(* Logix 5000 project; controller MV vendor 1 type 14 code 217 rev 31.11; software revision 31.00; part 24 of 53 *)
(* tags used below, declared in another part *)
   CheckTimeMask : INT;
   CWD : CHECKWORD_FLAGS;
   Delphi_Does_Eng_Func : BOOL;
   MC_CH1_FM_AI : PlantItem;   // CH1_FM
   MC_CH1_PTX_AI : PlantItem;   // CH1_PTX
   MC_CH2_FM_AI : PlantItem;   // CH2_FM
   MC_CH2_PTX_AI : PlantItem;   // CH2_PTX
   MC_CIP_AV09 : PlantItem;   // CIP_AV09
   MC_N100 : INT[255];   // C1_PLC Channel 1 PLC data
   MC_N100_29_1_Storagebit : BOOL;
   MC_N100_29_2_Storagebit : BOOL;
   MC_N100_29_3_Storagebit : BOOL;
   MC_N100_29_4_Storagebit : BOOL;
   MC_N102 : INT[255];   // CH1 PROG Channel 1 CIP progra m
   MC_N120 : INT[255];   // C2 PLC Channel 2 PLC data
   MC_N120_29_1_Storagebit : BOOL;
   MC_N120_29_2_Storagebit : BOOL;
   MC_N120_29_3_Storagebit : BOOL;
   MC_N120_29_4_Storagebit : BOOL;
   MC_N122 : INT[255];   // CH2 PROG Channel 2 CIP progra m
   MC_N20 : INT[255];   // P1 PRESS Control block and da ta for P1 pressure P ID loop
   MC_N21 : INT[255];   // P1 FLOW Control block and da ta for P1 flowrate P ID loop
   MC_N22 : INT[255];   // P2 PRESS Control block and da ta for P2 pressure P ID loop
   MC_N23 : INT[255];   // P2 FLOW Control block and da ta for P2 flowrate P ID loop
   MC_N255 : INT[255];   // CHECKWORDS Plant item checkword s
   MC_P1 : PlantItem;   // P1
   MC_P1_Flow_PID : PID;
   MC_P1_Flow_PID_Output : REAL;
   MC_P1_Pressure_PID : PID;
   MC_P1_Pressure_PID_Output : REAL;
   MC_P1_SP_AO : PlantItem;   // P1_SP
   MC_P2 : PlantItem;   // P2
   MC_P2_Flow_PID : PID;
   MC_P2_Flow_PID_Output : REAL;
   MC_P2_Pressure_PID : PID;
   MC_P2_Pressure_PID_Output : REAL;
   MC_P2_SP_AO : PlantItem;   // P2_SP
   TempChecktime : DINT;
(* MC_Common, continued *)

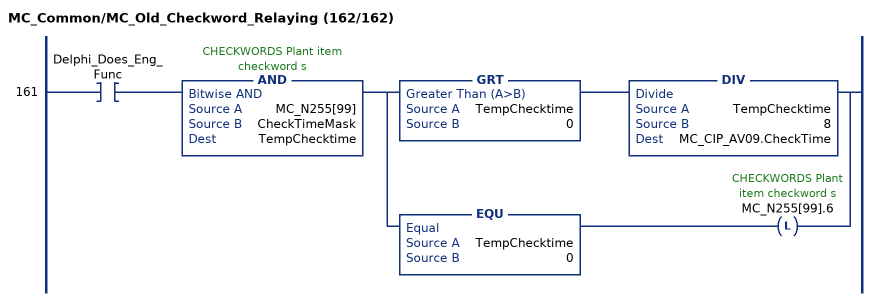
   [picture p434: MC_Common/MC_Old_Checkword_Relaying rungs 161-161]
   161: XIC(Delphi_Does_Eng_Func)AND(MC_N255[99],CheckTimeMask,TempChecktime)[GRT(TempChecktime,0) DIV(TempChecktime,8,MC_CIP_AV09.CheckTime) ,EQU(TempChecktime,0) OTL(MC_N255[99].6) ];
END_ROUTINE

ROUTINE MC_P1_FLOW_21   (* ladder *)
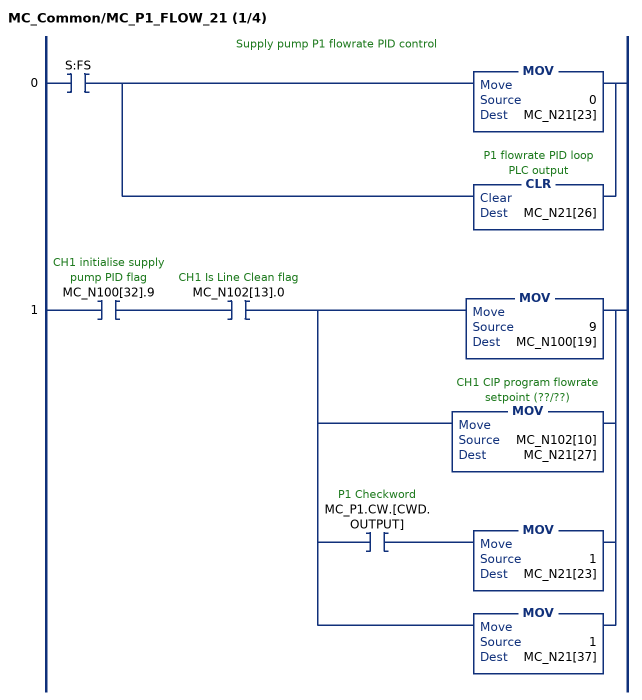
   // Supply pump P1 flowrate PID control
   0: XIC(S:FS)[MOV(0,MC_N21[23]) ,CLR(MC_N21[26]) ];
   1: XIC(MC_N100[32].9)XIC(MC_N102[13].0)[MOV(9,MC_N100[19]) ,MOV(MC_N102[10],MC_N21[27]) ,XIC(MC_P1.CW.[CWD.OUTPUT]) MOV(1,MC_N21[23]) ,MOV(1,MC_N21[37]) ];
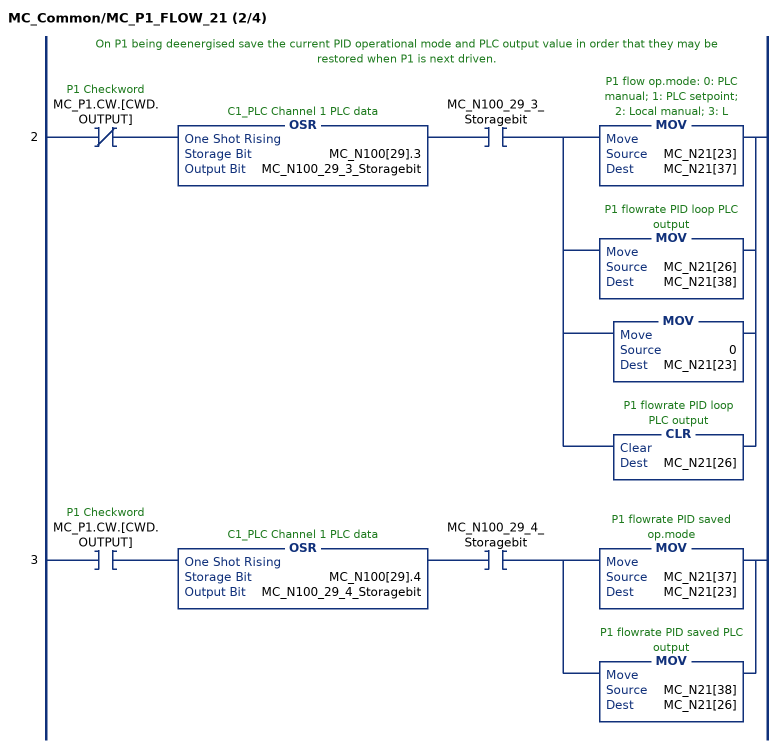
   // On P1 being deenergised save the current PID operational mode and PLC output value in order that they may be restored when P1 is next driven.
   2: XIO(MC_P1.CW.[CWD.OUTPUT])OSR(MC_N100[29].3,MC_N100_29_3_Storagebit)XIC(MC_N100_29_3_Storagebit)[MOV(MC_N21[23],MC_N21[37]) ,MOV(MC_N21[26],MC_N21[38]) ,MOV(0,MC_N21[23]) ,CLR(MC_N21[26]) ];
   3: XIC(MC_P1.CW.[CWD.OUTPUT])OSR(MC_N100[29].4,MC_N100_29_4_Storagebit)XIC(MC_N100_29_4_Storagebit)[MOV(MC_N21[37],MC_N21[23]) ,MOV(MC_N21[38],MC_N21[26]) ];
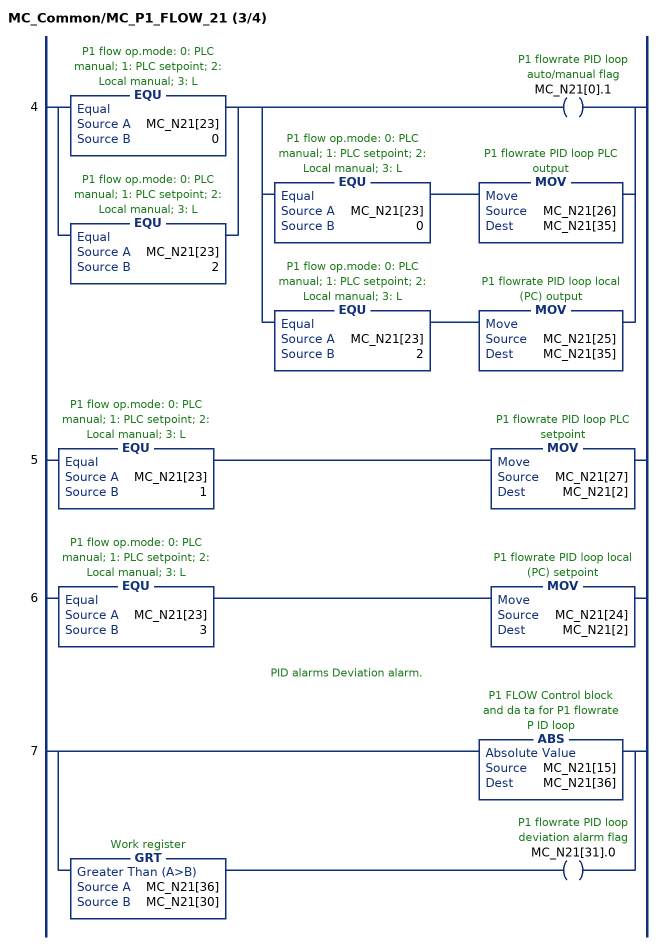
   4: [EQU(MC_N21[23],0) ,EQU(MC_N21[23],2) ][OTE(MC_N21[0].1) ,EQU(MC_N21[23],0) MOV(MC_N21[26],MC_N21[35]) ,EQU(MC_N21[23],2) MOV(MC_N21[25],MC_N21[35]) ];
   5: EQU(MC_N21[23],1)MOV(MC_N21[27],MC_N21[2]);
   6: EQU(MC_N21[23],3)MOV(MC_N21[24],MC_N21[2]);
   // PID alarms Deviation alarm.
   7: [ABS(MC_N21[15],MC_N21[36]) ,GRT(MC_N21[36],MC_N21[30]) OTE(MC_N21[31].0) ];
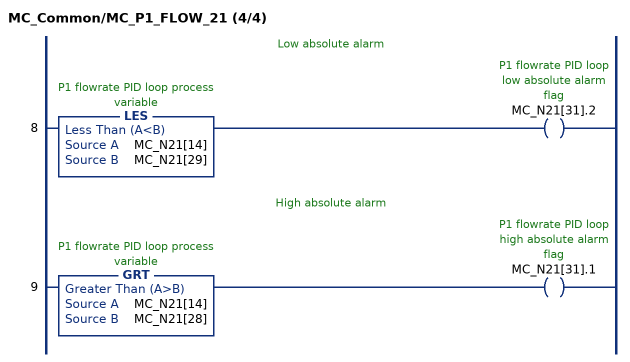
   // Low absolute alarm
   8: LES(MC_N21[14],MC_N21[29])OTE(MC_N21[31].2);
   // High absolute alarm
   9: GRT(MC_N21[14],MC_N21[28])OTE(MC_N21[31].1);
END_ROUTINE

ROUTINE MC_P1_PRESS_20   (* ladder *)
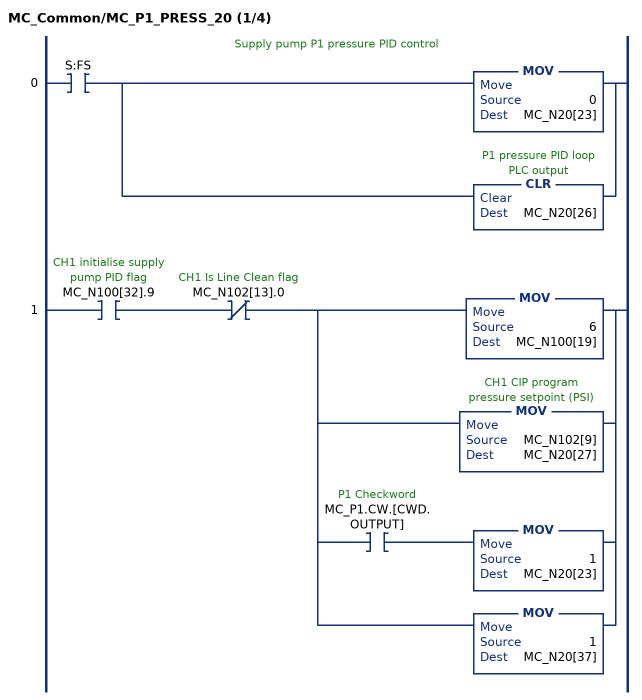
   // Supply pump P1 pressure PID control
   0: XIC(S:FS)[MOV(0,MC_N20[23]) ,CLR(MC_N20[26]) ];
   1: XIC(MC_N100[32].9)XIO(MC_N102[13].0)[MOV(6,MC_N100[19]) ,MOV(MC_N102[9],MC_N20[27]) ,XIC(MC_P1.CW.[CWD.OUTPUT]) MOV(1,MC_N20[23]) ,MOV(1,MC_N20[37]) ];
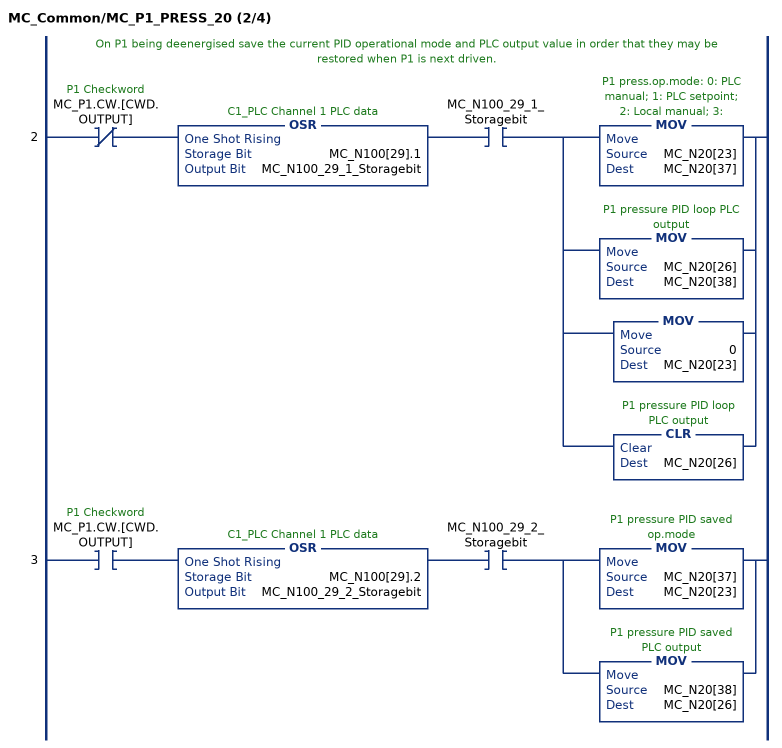
   // On P1 being deenergised save the current PID operational mode and PLC output value in order that they may be restored when P1 is next driven.
   2: XIO(MC_P1.CW.[CWD.OUTPUT])OSR(MC_N100[29].1,MC_N100_29_1_Storagebit)XIC(MC_N100_29_1_Storagebit)[MOV(MC_N20[23],MC_N20[37]) ,MOV(MC_N20[26],MC_N20[38]) ,MOV(0,MC_N20[23]) ,CLR(MC_N20[26]) ];
   3: XIC(MC_P1.CW.[CWD.OUTPUT])OSR(MC_N100[29].2,MC_N100_29_2_Storagebit)XIC(MC_N100_29_2_Storagebit)[MOV(MC_N20[37],MC_N20[23]) ,MOV(MC_N20[38],MC_N20[26]) ];
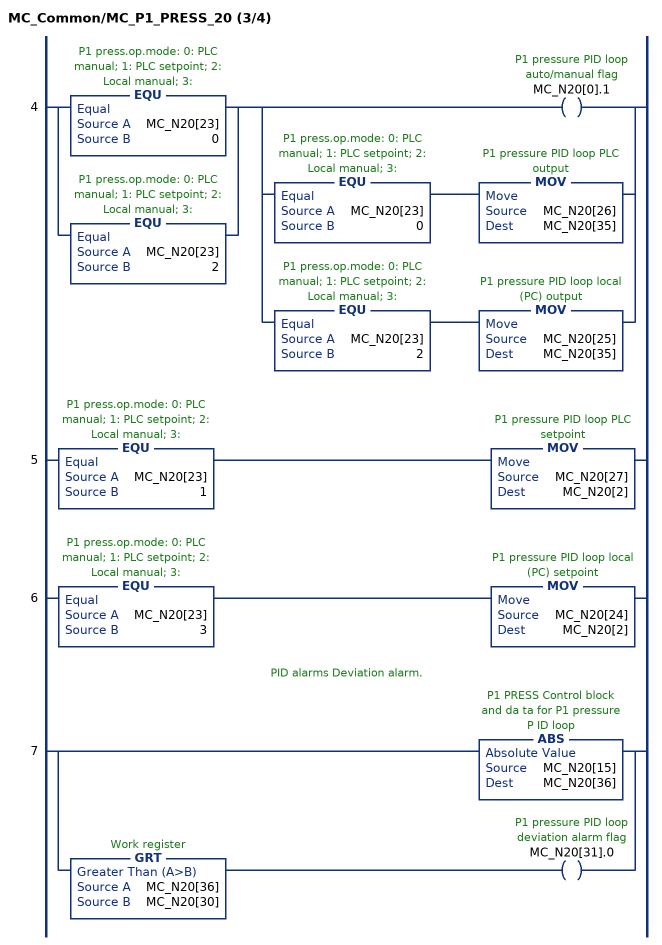
   4: [EQU(MC_N20[23],0) ,EQU(MC_N20[23],2) ][OTE(MC_N20[0].1) ,EQU(MC_N20[23],0) MOV(MC_N20[26],MC_N20[35]) ,EQU(MC_N20[23],2) MOV(MC_N20[25],MC_N20[35]) ];
   5: EQU(MC_N20[23],1)MOV(MC_N20[27],MC_N20[2]);
   6: EQU(MC_N20[23],3)MOV(MC_N20[24],MC_N20[2]);
   // PID alarms Deviation alarm.
   7: [ABS(MC_N20[15],MC_N20[36]) ,GRT(MC_N20[36],MC_N20[30]) OTE(MC_N20[31].0) ];
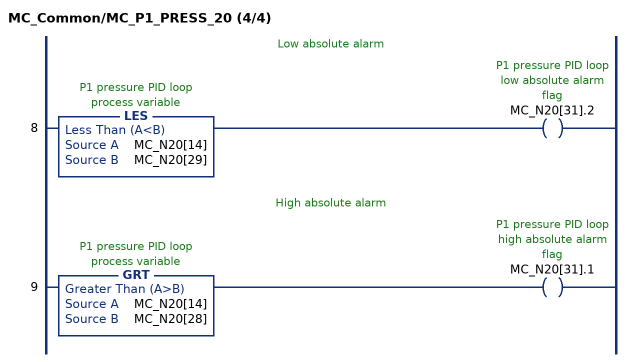
   // Low absolute alarm
   8: LES(MC_N20[14],MC_N20[29])OTE(MC_N20[31].2);
   // High absolute alarm
   9: GRT(MC_N20[14],MC_N20[28])OTE(MC_N20[31].1);
END_ROUTINE

ROUTINE MC_P2_FLOW_23   (* ladder *)
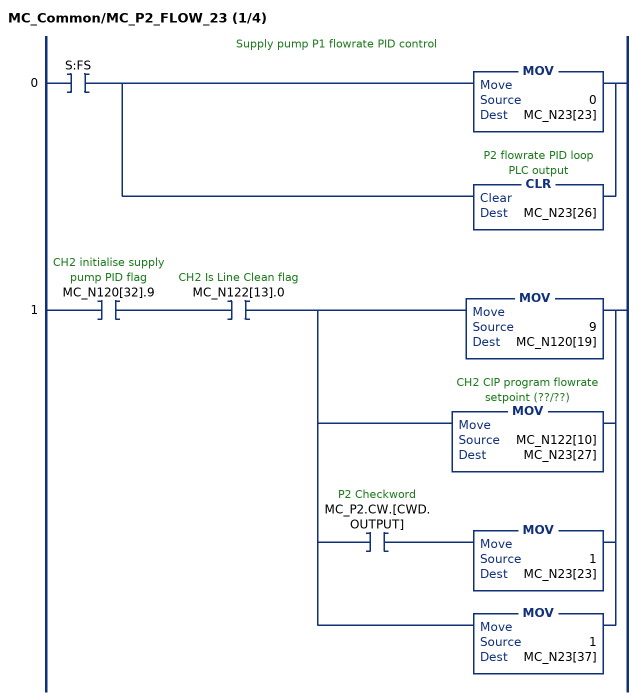
   // Supply pump P1 flowrate PID control
   0: XIC(S:FS)[MOV(0,MC_N23[23]) ,CLR(MC_N23[26]) ];
   1: XIC(MC_N120[32].9)XIC(MC_N122[13].0)[MOV(9,MC_N120[19]) ,MOV(MC_N122[10],MC_N23[27]) ,XIC(MC_P2.CW.[CWD.OUTPUT]) MOV(1,MC_N23[23]) ,MOV(1,MC_N23[37]) ];
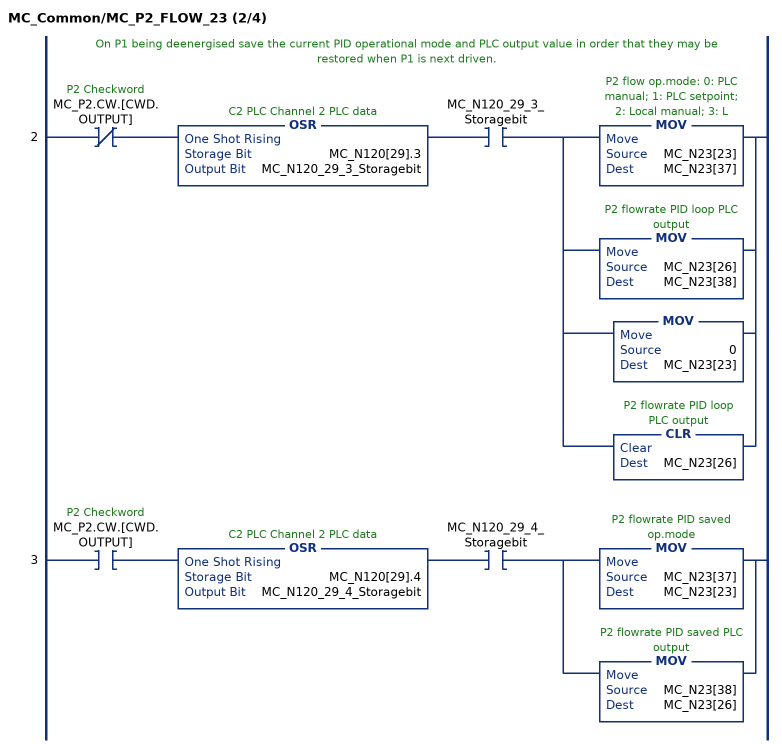
   // On P1 being deenergised save the current PID operational mode and PLC output value in order that they may be restored when P1 is next driven.
   2: XIO(MC_P2.CW.[CWD.OUTPUT])OSR(MC_N120[29].3,MC_N120_29_3_Storagebit)XIC(MC_N120_29_3_Storagebit)[MOV(MC_N23[23],MC_N23[37]) ,MOV(MC_N23[26],MC_N23[38]) ,MOV(0,MC_N23[23]) ,CLR(MC_N23[26]) ];
   3: XIC(MC_P2.CW.[CWD.OUTPUT])OSR(MC_N120[29].4,MC_N120_29_4_Storagebit)XIC(MC_N120_29_4_Storagebit)[MOV(MC_N23[37],MC_N23[23]) ,MOV(MC_N23[38],MC_N23[26]) ];
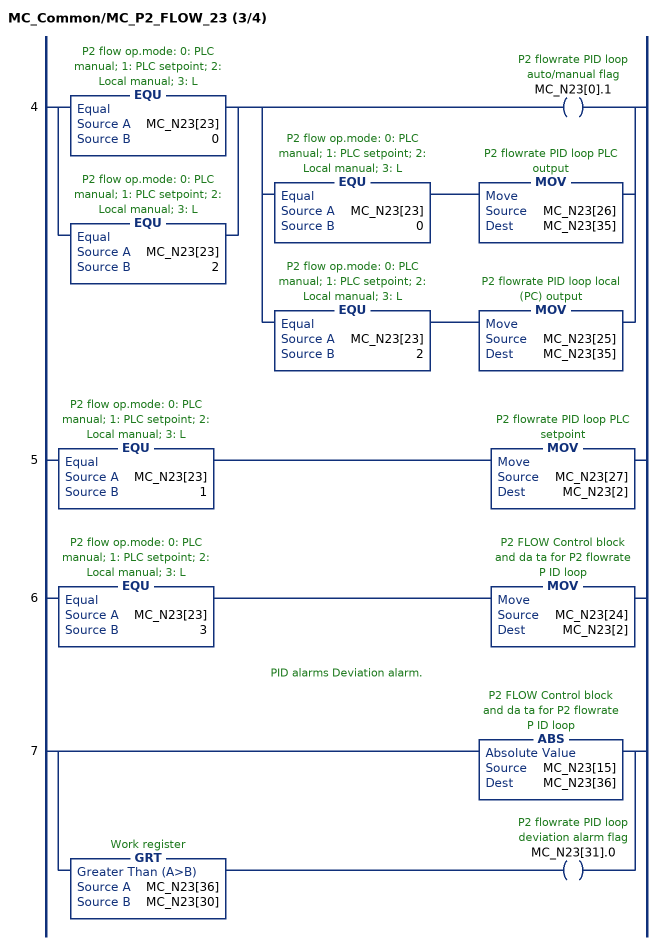
   4: [EQU(MC_N23[23],0) ,EQU(MC_N23[23],2) ][OTE(MC_N23[0].1) ,EQU(MC_N23[23],0) MOV(MC_N23[26],MC_N23[35]) ,EQU(MC_N23[23],2) MOV(MC_N23[25],MC_N23[35]) ];
   5: EQU(MC_N23[23],1)MOV(MC_N23[27],MC_N23[2]);
   6: EQU(MC_N23[23],3)MOV(MC_N23[24],MC_N23[2]);
   // PID alarms Deviation alarm.
   7: [ABS(MC_N23[15],MC_N23[36]) ,GRT(MC_N23[36],MC_N23[30]) OTE(MC_N23[31].0) ];
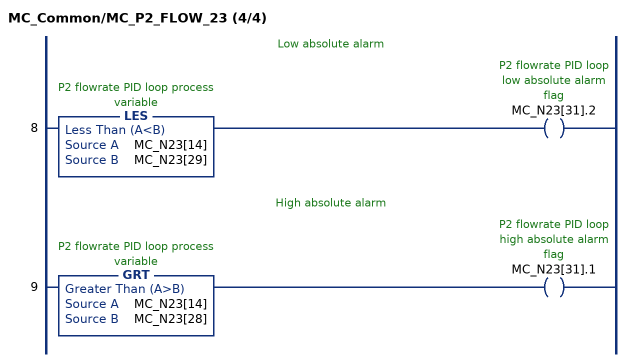
   // Low absolute alarm
   8: LES(MC_N23[14],MC_N23[29])OTE(MC_N23[31].2);
   // High absolute alarm
   9: GRT(MC_N23[14],MC_N23[28])OTE(MC_N23[31].1);
END_ROUTINE

ROUTINE MC_P2_PRESS_22   (* ladder *)
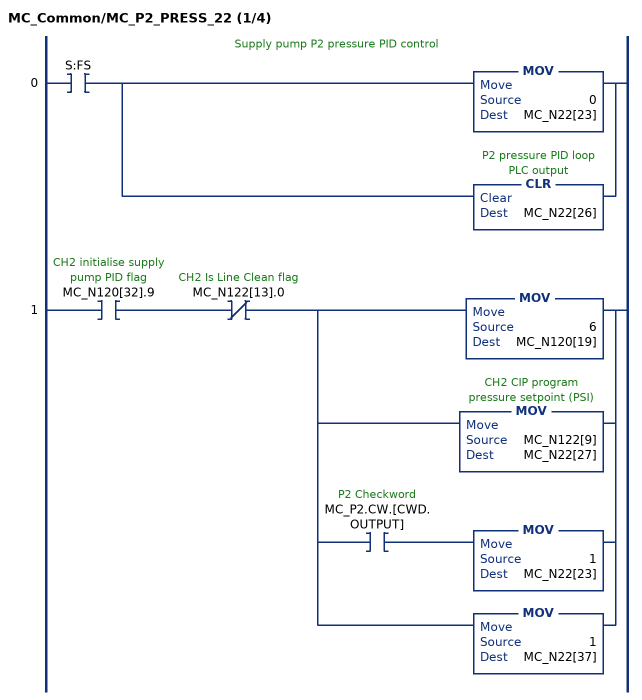
   // Supply pump P2 pressure PID control
   0: XIC(S:FS)[MOV(0,MC_N22[23]) ,CLR(MC_N22[26]) ];
   1: XIC(MC_N120[32].9)XIO(MC_N122[13].0)[MOV(6,MC_N120[19]) ,MOV(MC_N122[9],MC_N22[27]) ,XIC(MC_P2.CW.[CWD.OUTPUT]) MOV(1,MC_N22[23]) ,MOV(1,MC_N22[37]) ];
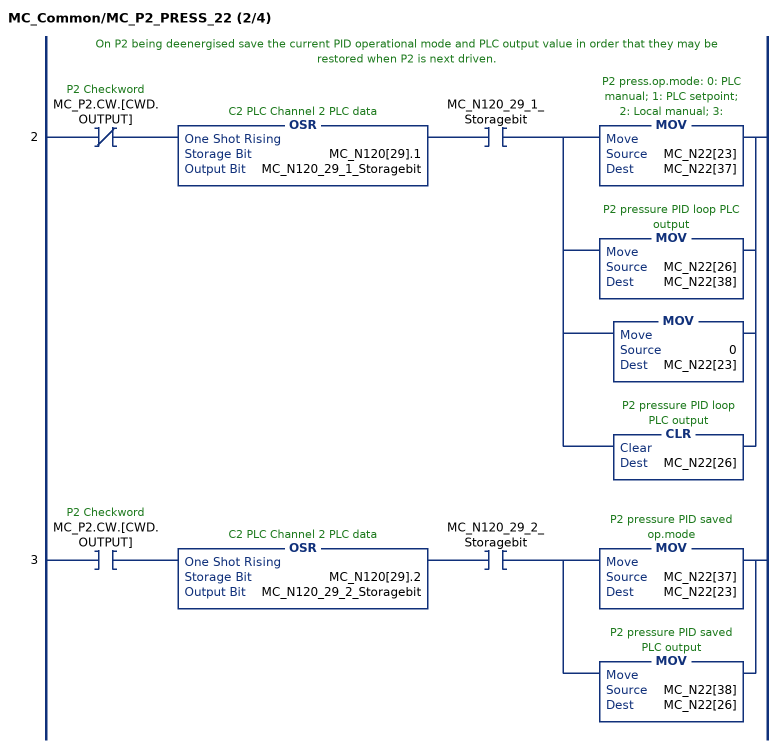
   // On P2 being deenergised save the current PID operational mode and PLC output value in order that they may be restored when P2 is next driven.
   2: XIO(MC_P2.CW.[CWD.OUTPUT])OSR(MC_N120[29].1,MC_N120_29_1_Storagebit)XIC(MC_N120_29_1_Storagebit)[MOV(MC_N22[23],MC_N22[37]) ,MOV(MC_N22[26],MC_N22[38]) ,MOV(0,MC_N22[23]) ,CLR(MC_N22[26]) ];
   3: XIC(MC_P2.CW.[CWD.OUTPUT])OSR(MC_N120[29].2,MC_N120_29_2_Storagebit)XIC(MC_N120_29_2_Storagebit)[MOV(MC_N22[37],MC_N22[23]) ,MOV(MC_N22[38],MC_N22[26]) ];
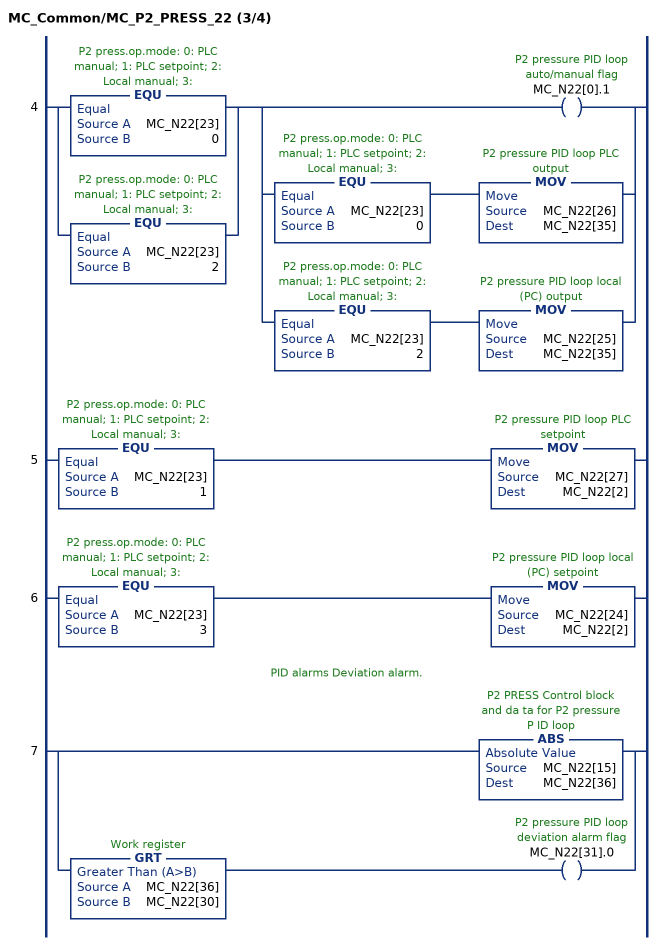
   4: [EQU(MC_N22[23],0) ,EQU(MC_N22[23],2) ][OTE(MC_N22[0].1) ,EQU(MC_N22[23],0) MOV(MC_N22[26],MC_N22[35]) ,EQU(MC_N22[23],2) MOV(MC_N22[25],MC_N22[35]) ];
   5: EQU(MC_N22[23],1)MOV(MC_N22[27],MC_N22[2]);
   6: EQU(MC_N22[23],3)MOV(MC_N22[24],MC_N22[2]);
   // PID alarms Deviation alarm.
   7: [ABS(MC_N22[15],MC_N22[36]) ,GRT(MC_N22[36],MC_N22[30]) OTE(MC_N22[31].0) ];
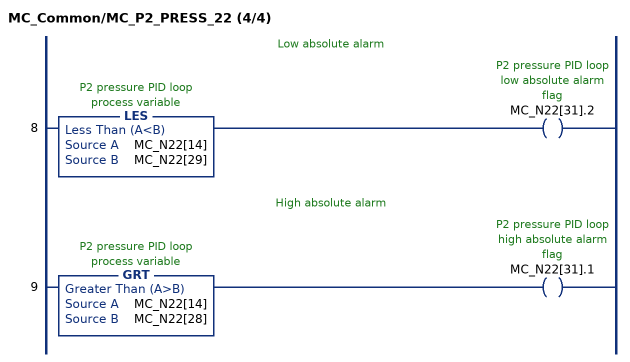
   // Low absolute alarm
   8: LES(MC_N22[14],MC_N22[29])OTE(MC_N22[31].2);
   // High absolute alarm
   9: GRT(MC_N22[14],MC_N22[28])OTE(MC_N22[31].1);
END_ROUTINE

ROUTINE MC_PID_18   (* ladder *)
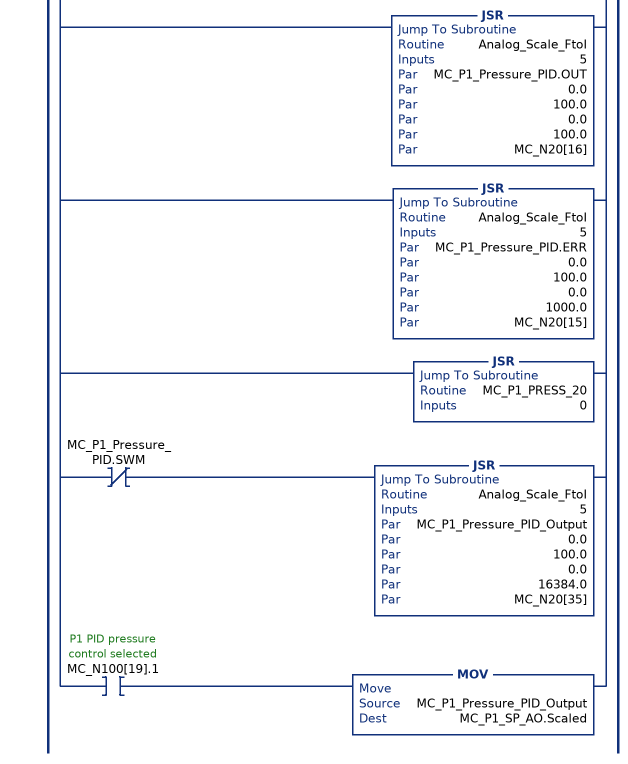
   // PID controllers Channel 1(pump P1) pressure control
   0: [XIC(MC_N20[0].1) OTE(MC_P1_Pressure_PID.SWM) ,JSR(Analog_Scale_ItoF,5,MC_N20[2],0.0,1000.0,0.0,100.0,MC_P1_Pressure_PID.SP) ,JSR(Analog_Scale_FtoI,5,MC_CH1_PTX_AI.Scaled,0.0,100.0,0.0,16384.0,MC_N20[34]) ,XIC(MC_P1_Pressure_PID.SWM) JSR(Analog_Scale_ItoF,5,MC_N20[35],0.0,16384.0,0.0,100.0,MC_P1_Pressure_PID.SO) ,PID(MC_P1_Pressure_PID,MC_CH1_PTX_AI.Scaled,MC_P1_Pressure_PID_Output,MC_P1_Pressure_PID_Output,0,0,0) ,JSR(Analog_Scale_FtoI,5,MC_P1_Pressure_PID.PV,0.0,100.0,0.0,1000.0,MC_N20[14]) ,JSR(Analog_Scale_FtoI,5,MC_P1_Pressure_PID.OUT,0.0,100.0,0.0,100.0,MC_N20[16]) ,JSR(Analog_Scale_FtoI,5,MC_P1_Pressure_PID.ERR,0.0,100.0,0.0,1000.0,MC_N20[15]) ,JSR(MC_P1_PRESS_20,0) ,XIO(MC_P1_Pressure_PID.SWM) JSR(Analog_Scale_FtoI,5,MC_P1_Pressure_PID_Output,0.0,100.0,0.0,16384.0,MC_N20[35]) ,XIC(MC_N100[19].1) MOV(MC_P1_Pressure_PID_Output,MC_P1_SP_AO.Scaled) ];
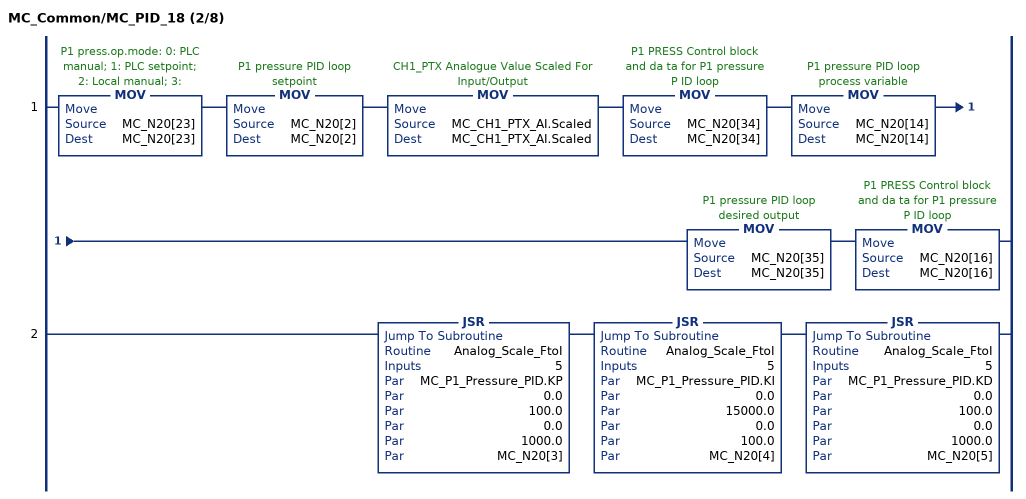
   1: MOV(MC_N20[23],MC_N20[23])MOV(MC_N20[2],MC_N20[2])MOV(MC_CH1_PTX_AI.Scaled,MC_CH1_PTX_AI.Scaled)MOV(MC_N20[34],MC_N20[34])MOV(MC_N20[14],MC_N20[14])MOV(MC_N20[35],MC_N20[35])MOV(MC_N20[16],MC_N20[16]);
   2: JSR(Analog_Scale_FtoI,5,MC_P1_Pressure_PID.KP,0.0,100.0,0.0,1000.0,MC_N20[3])JSR(Analog_Scale_FtoI,5,MC_P1_Pressure_PID.KI,0.0,15000.0,0.0,100.0,MC_N20[4])JSR(Analog_Scale_FtoI,5,MC_P1_Pressure_PID.KD,0.0,100.0,0.0,1000.0,MC_N20[5]);
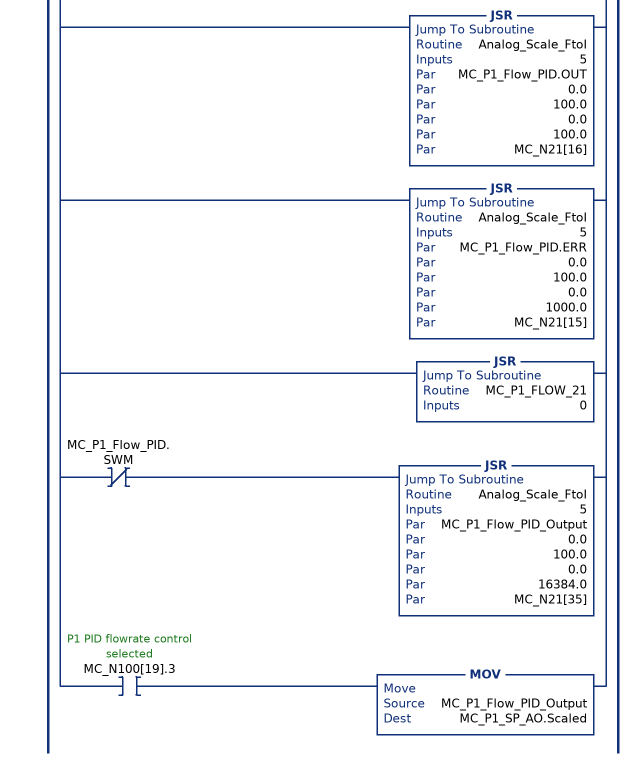
   // Channel 1 (pump P1) flowrate control
   3: [XIC(MC_N21[0].1) OTE(MC_P1_Flow_PID.SWM) ,JSR(Analog_Scale_ItoF,5,MC_N21[2],0.0,1000.0,0.0,100.0,MC_P1_Flow_PID.SP) ,JSR(Analog_Scale_FtoI,5,MC_CH1_FM_AI.Scaled,0.0,500.0,0.0,16384.0,MC_N21[34]) ,XIC(MC_P1_Flow_PID.SWM) JSR(Analog_Scale_ItoF,5,MC_N21[35],0.0,16384.0,0.0,100.0,MC_P1_Flow_PID.SO) ,PID(MC_P1_Flow_PID,MC_CH1_FM_AI.Scaled,MC_P1_Flow_PID_Output,MC_P1_Flow_PID_Output,0,0,0) ,JSR(Analog_Scale_FtoI,5,MC_P1_Flow_PID.PV,0.0,100.0,0.0,1000.0,MC_N21[14]) ,JSR(Analog_Scale_FtoI,5,MC_P1_Flow_PID.OUT,0.0,100.0,0.0,100.0,MC_N21[16]) ,JSR(Analog_Scale_FtoI,5,MC_P1_Flow_PID.ERR,0.0,100.0,0.0,1000.0,MC_N21[15]) ,JSR(MC_P1_FLOW_21,0) ,XIO(MC_P1_Flow_PID.SWM) JSR(Analog_Scale_FtoI,5,MC_P1_Flow_PID_Output,0.0,100.0,0.0,16384.0,MC_N21[35]) ,XIC(MC_N100[19].3) MOV(MC_P1_Flow_PID_Output,MC_P1_SP_AO.Scaled) ];
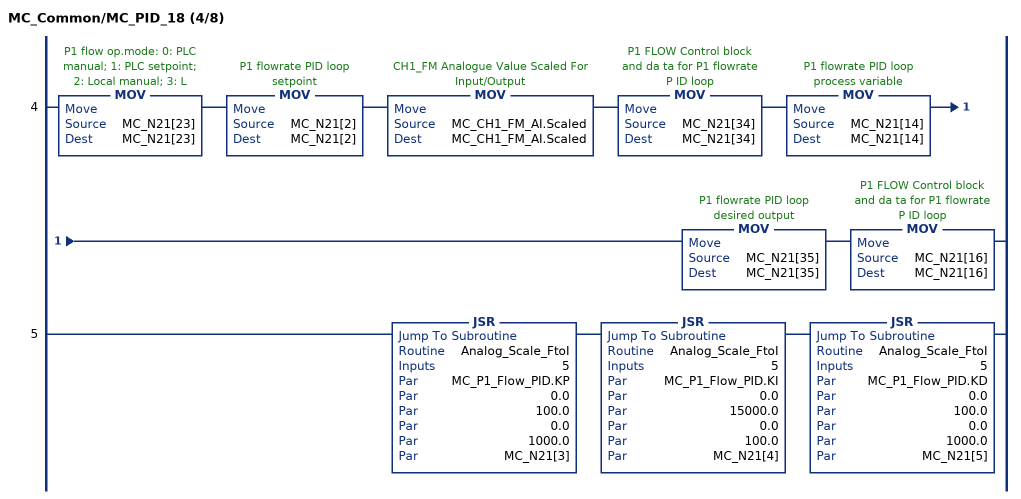
   4: MOV(MC_N21[23],MC_N21[23])MOV(MC_N21[2],MC_N21[2])MOV(MC_CH1_FM_AI.Scaled,MC_CH1_FM_AI.Scaled)MOV(MC_N21[34],MC_N21[34])MOV(MC_N21[14],MC_N21[14])MOV(MC_N21[35],MC_N21[35])MOV(MC_N21[16],MC_N21[16]);
   5: JSR(Analog_Scale_FtoI,5,MC_P1_Flow_PID.KP,0.0,100.0,0.0,1000.0,MC_N21[3])JSR(Analog_Scale_FtoI,5,MC_P1_Flow_PID.KI,0.0,15000.0,0.0,100.0,MC_N21[4])JSR(Analog_Scale_FtoI,5,MC_P1_Flow_PID.KD,0.0,100.0,0.0,1000.0,MC_N21[5]);
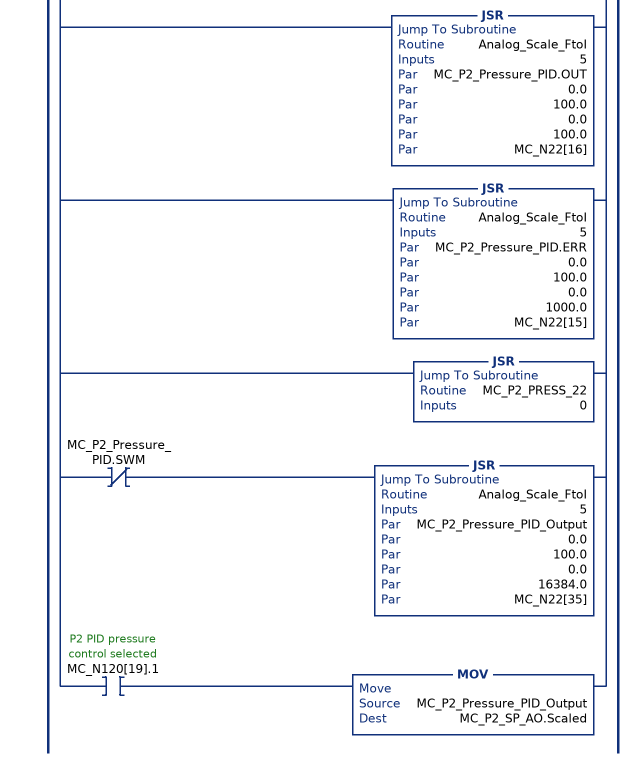
   // Channel 2 (pump P2) pressure control
   6: [XIC(MC_N22[0].1) OTE(MC_P2_Pressure_PID.SWM) ,JSR(Analog_Scale_ItoF,5,MC_N22[2],0.0,1000.0,0.0,100.0,MC_P2_Pressure_PID.SP) ,JSR(Analog_Scale_FtoI,5,MC_CH2_PTX_AI.Scaled,0.0,100.0,0.0,16384.0,MC_N22[34]) ,XIC(MC_P2_Pressure_PID.SWM) JSR(Analog_Scale_ItoF,5,MC_N22[35],0.0,16384.0,0.0,100.0,MC_P2_Pressure_PID.SO) ,PID(MC_P2_Pressure_PID,MC_CH2_PTX_AI.Scaled,MC_P2_Pressure_PID_Output,MC_P2_Pressure_PID_Output,0,0,0) ,JSR(Analog_Scale_FtoI,5,MC_P2_Pressure_PID.PV,0.0,100.0,0.0,1000.0,MC_N22[14]) ,JSR(Analog_Scale_FtoI,5,MC_P2_Pressure_PID.OUT,0.0,100.0,0.0,100.0,MC_N22[16]) ,JSR(Analog_Scale_FtoI,5,MC_P2_Pressure_PID.ERR,0.0,100.0,0.0,1000.0,MC_N22[15]) ,JSR(MC_P2_PRESS_22,0) ,XIO(MC_P2_Pressure_PID.SWM) JSR(Analog_Scale_FtoI,5,MC_P2_Pressure_PID_Output,0.0,100.0,0.0,16384.0,MC_N22[35]) ,XIC(MC_N120[19].1) MOV(MC_P2_Pressure_PID_Output,MC_P2_SP_AO.Scaled) ];
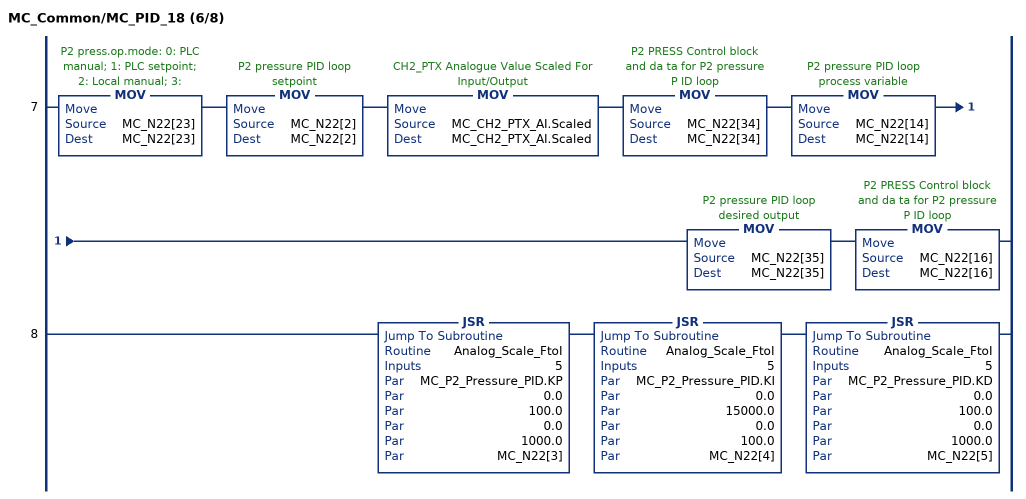
   7: MOV(MC_N22[23],MC_N22[23])MOV(MC_N22[2],MC_N22[2])MOV(MC_CH2_PTX_AI.Scaled,MC_CH2_PTX_AI.Scaled)MOV(MC_N22[34],MC_N22[34])MOV(MC_N22[14],MC_N22[14])MOV(MC_N22[35],MC_N22[35])MOV(MC_N22[16],MC_N22[16]);
   8: JSR(Analog_Scale_FtoI,5,MC_P2_Pressure_PID.KP,0.0,100.0,0.0,1000.0,MC_N22[3])JSR(Analog_Scale_FtoI,5,MC_P2_Pressure_PID.KI,0.0,15000.0,0.0,100.0,MC_N22[4])JSR(Analog_Scale_FtoI,5,MC_P2_Pressure_PID.KD,0.0,100.0,0.0,1000.0,MC_N22[5]);
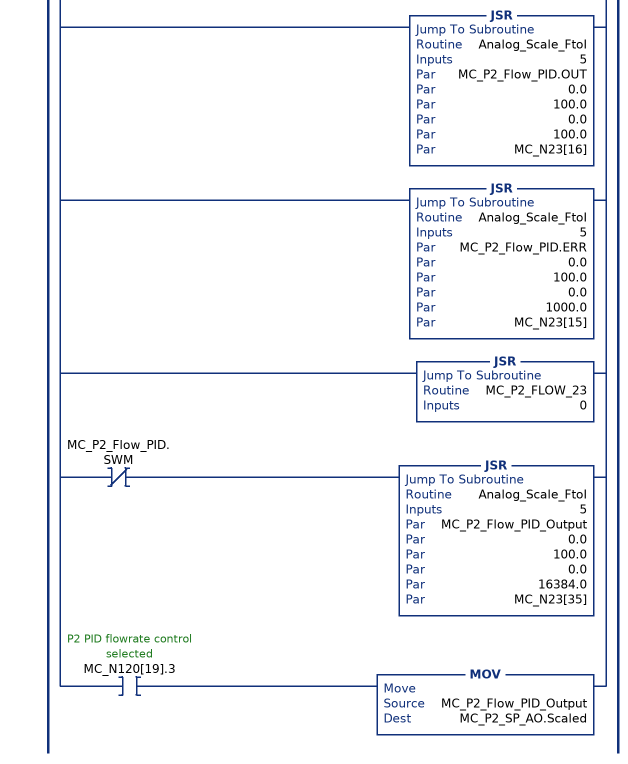
   // Channel 2 (pump P2) flowrate control
   9: [XIC(MC_N23[0].1) OTE(MC_P2_Flow_PID.SWM) ,JSR(Analog_Scale_ItoF,5,MC_N23[2],0.0,1000.0,0.0,100.0,MC_P2_Flow_PID.SP) ,JSR(Analog_Scale_FtoI,5,MC_CH2_FM_AI.Scaled,0.0,500.0,0.0,16384.0,MC_N23[34]) ,XIC(MC_P2_Flow_PID.SWM) JSR(Analog_Scale_ItoF,5,MC_N23[35],0.0,16384.0,0.0,100.0,MC_P2_Flow_PID.SO) ,PID(MC_P2_Flow_PID,MC_CH2_FM_AI.Scaled,MC_P2_Flow_PID_Output,MC_P2_Flow_PID_Output,0,0,0) ,JSR(Analog_Scale_FtoI,5,MC_P2_Flow_PID.PV,0.0,100.0,0.0,1000.0,MC_N23[14]) ,JSR(Analog_Scale_FtoI,5,MC_P2_Flow_PID.OUT,0.0,100.0,0.0,100.0,MC_N23[16]) ,JSR(Analog_Scale_FtoI,5,MC_P2_Flow_PID.ERR,0.0,100.0,0.0,1000.0,MC_N23[15]) ,JSR(MC_P2_FLOW_23,0) ,XIO(MC_P2_Flow_PID.SWM) JSR(Analog_Scale_FtoI,5,MC_P2_Flow_PID_Output,0.0,100.0,0.0,16384.0,MC_N23[35]) ,XIC(MC_N120[19].3) MOV(MC_P2_Flow_PID_Output,MC_P2_SP_AO.Scaled) ];
